(* Logix 5000 project; controller OWF Emulate 5570 rev 30.12; software revision 30.00; part 18 of 21 *)
(* tags used below, declared in another part *)
   OWF_Add_c : DINT;
   OWF_Input : DINT[16];
   OWF_Result : DINT[17];
(* MainProgram, continued *)

   		OWF_Result[4].31:=0;
   		OWF_Result[5]:=OWF_Result[5] + 1895099717+OWF_Add_c;
   		OWF_Add_c.5:=OWF_Result[5].31;
   		OWF_Result[5].31:=0;
   		OWF_Result[6]:=OWF_Result[6] + 2009701654+OWF_Add_c;
   		OWF_Add_c.6:=OWF_Result[6].31;
   		OWF_Result[6].31:=0;
   		OWF_Result[7]:=OWF_Result[7] + 1963030177+OWF_Add_c;
   		OWF_Add_c.7:=OWF_Result[7].31;
   		OWF_Result[7].31:=0;
   		OWF_Result[8]:=OWF_Result[8] + 232130595+OWF_Add_c;
   		OWF_Add_c.8:=OWF_Result[8].31;
   		OWF_Result[8].31:=0;
   		OWF_Result[9]:=OWF_Result[9] + 1484597708+OWF_Add_c;
   		OWF_Add_c.9:=OWF_Result[9].31;
   		OWF_Result[9].31:=0;
   		OWF_Result[10]:=OWF_Result[10] + 955822561+OWF_Add_c;
   		OWF_Add_c.10:=OWF_Result[10].31;
   		OWF_Result[10].31:=0;
   		OWF_Result[11]:=OWF_Result[11] + 760226904+OWF_Add_c;
   		OWF_Add_c.11:=OWF_Result[11].31;
   		OWF_Result[11].31:=0;
   		OWF_Result[12]:=OWF_Result[12] + 1637968730+OWF_Add_c;
   		OWF_Add_c.12:=OWF_Result[12].31;
   		OWF_Result[12].31:=0;
   		OWF_Result[13]:=OWF_Result[13] + 1060225387+OWF_Add_c;
   		OWF_Add_c.13:=OWF_Result[13].31;
   		OWF_Result[13].31:=0;
   		OWF_Result[14]:=OWF_Result[14] + 1695671309+OWF_Add_c;
   		OWF_Add_c.14:=OWF_Result[14].31;
   		OWF_Result[14].31:=0;
   		OWF_Result[15]:=OWF_Result[15] + 2141154184+OWF_Add_c;
   		OWF_Add_c.15:=OWF_Result[15].31;
   		OWF_Result[15].31:=0;
   		OWF_Result[16]:=OWF_Result[16] + 1403333060+OWF_Add_c;
   		OWF_Add_c.16:=OWF_Result[16].31;
   		OWF_Result[16].31:=0;
   	End_If;
   	If OWF_Input[11].[13] Then
   		OWF_Result[0]:=OWF_Result[0] + 1424989119+OWF_Add_c;
   		OWF_Add_c.0:=OWF_Result[0].31;
   		OWF_Result[0].31:=0;
   		OWF_Result[1]:=OWF_Result[1] + 1792831216+OWF_Add_c;
   		OWF_Add_c.1:=OWF_Result[1].31;
   		OWF_Result[1].31:=0;
   		OWF_Result[2]:=OWF_Result[2] + 1280480339+OWF_Add_c;
   		OWF_Add_c.2:=OWF_Result[2].31;
   		OWF_Result[2].31:=0;
   		OWF_Result[3]:=OWF_Result[3] + 1887620187+OWF_Add_c;
   		OWF_Add_c.3:=OWF_Result[3].31;
   		OWF_Result[3].31:=0;
   		OWF_Result[4]:=OWF_Result[4] + 50882950+OWF_Add_c;
   		OWF_Add_c.4:=OWF_Result[4].31;
   		OWF_Result[4].31:=0;
   		OWF_Result[5]:=OWF_Result[5] + 1542129432+OWF_Add_c;
   		OWF_Add_c.5:=OWF_Result[5].31;
   		OWF_Result[5].31:=0;
   		OWF_Result[6]:=OWF_Result[6] + 1234316724+OWF_Add_c;
   		OWF_Add_c.6:=OWF_Result[6].31;
   		OWF_Result[6].31:=0;
   		OWF_Result[7]:=OWF_Result[7] + 267891254+OWF_Add_c;
   		OWF_Add_c.7:=OWF_Result[7].31;
   		OWF_Result[7].31:=0;
   		OWF_Result[8]:=OWF_Result[8] + 1066053149+OWF_Add_c;
   		OWF_Add_c.8:=OWF_Result[8].31;
   		OWF_Result[8].31:=0;
   		OWF_Result[9]:=OWF_Result[9] + 54187296+OWF_Add_c;
   		OWF_Add_c.9:=OWF_Result[9].31;
   		OWF_Result[9].31:=0;
   		OWF_Result[10]:=OWF_Result[10] + 129651269+OWF_Add_c;
   		OWF_Add_c.10:=OWF_Result[10].31;
   		OWF_Result[10].31:=0;
   		OWF_Result[11]:=OWF_Result[11] + 604389954+OWF_Add_c;
   		OWF_Add_c.11:=OWF_Result[11].31;
   		OWF_Result[11].31:=0;
   		OWF_Result[12]:=OWF_Result[12] + 1474729667+OWF_Add_c;
   		OWF_Add_c.12:=OWF_Result[12].31;
   		OWF_Result[12].31:=0;
   		OWF_Result[13]:=OWF_Result[13] + 627513733+OWF_Add_c;
   		OWF_Add_c.13:=OWF_Result[13].31;
   		OWF_Result[13].31:=0;
   		OWF_Result[14]:=OWF_Result[14] + 1221285509+OWF_Add_c;
   		OWF_Add_c.14:=OWF_Result[14].31;
   		OWF_Result[14].31:=0;
   		OWF_Result[15]:=OWF_Result[15] + 1347886424+OWF_Add_c;
   		OWF_Add_c.15:=OWF_Result[15].31;
   		OWF_Result[15].31:=0;
   		OWF_Result[16]:=OWF_Result[16] + 1501741428+OWF_Add_c;
   		OWF_Add_c.16:=OWF_Result[16].31;
   		OWF_Result[16].31:=0;
   	End_If;
   	If OWF_Input[11].[14] Then
   		OWF_Result[0]:=OWF_Result[0] + 148251354+OWF_Add_c;
   		OWF_Add_c.0:=OWF_Result[0].31;
   		OWF_Result[0].31:=0;
   		OWF_Result[1]:=OWF_Result[1] + 734679875+OWF_Add_c;
   		OWF_Add_c.1:=OWF_Result[1].31;
   		OWF_Result[1].31:=0;
   		OWF_Result[2]:=OWF_Result[2] + 501019324+OWF_Add_c;
   		OWF_Add_c.2:=OWF_Result[2].31;
   		OWF_Result[2].31:=0;
   		OWF_Result[3]:=OWF_Result[3] + 1051894690+OWF_Add_c;
   		OWF_Add_c.3:=OWF_Result[3].31;
   		OWF_Result[3].31:=0;
   		OWF_Result[4]:=OWF_Result[4] + 713394787+OWF_Add_c;
   		OWF_Add_c.4:=OWF_Result[4].31;
   		OWF_Result[4].31:=0;
   		OWF_Result[5]:=OWF_Result[5] + 875122393+OWF_Add_c;
   		OWF_Add_c.5:=OWF_Result[5].31;
   		OWF_Result[5].31:=0;
   		OWF_Result[6]:=OWF_Result[6] + 259478417+OWF_Add_c;
   		OWF_Add_c.6:=OWF_Result[6].31;
   		OWF_Result[6].31:=0;
   		OWF_Result[7]:=OWF_Result[7] + 1855876414+OWF_Add_c;
   		OWF_Add_c.7:=OWF_Result[7].31;
   		OWF_Result[7].31:=0;
   		OWF_Result[8]:=OWF_Result[8] + 1892105+OWF_Add_c;
   		OWF_Add_c.8:=OWF_Result[8].31;
   		OWF_Result[8].31:=0;
   		OWF_Result[9]:=OWF_Result[9] + 229647947+OWF_Add_c;
   		OWF_Add_c.9:=OWF_Result[9].31;
   		OWF_Result[9].31:=0;
   		OWF_Result[10]:=OWF_Result[10] + 445153450+OWF_Add_c;
   		OWF_Add_c.10:=OWF_Result[10].31;
   		OWF_Result[10].31:=0;
   		OWF_Result[11]:=OWF_Result[11] + 1697696739+OWF_Add_c;
   		OWF_Add_c.11:=OWF_Result[11].31;
   		OWF_Result[11].31:=0;
   		OWF_Result[12]:=OWF_Result[12] + 259481221+OWF_Add_c;
   		OWF_Add_c.12:=OWF_Result[12].31;
   		OWF_Result[12].31:=0;
   		OWF_Result[13]:=OWF_Result[13] + 98481250+OWF_Add_c;
   		OWF_Add_c.13:=OWF_Result[13].31;
   		OWF_Result[13].31:=0;
   		OWF_Result[14]:=OWF_Result[14] + 6041701+OWF_Add_c;
   		OWF_Add_c.14:=OWF_Result[14].31;
   		OWF_Result[14].31:=0;
   		OWF_Result[15]:=OWF_Result[15] + 184524762+OWF_Add_c;
   		OWF_Add_c.15:=OWF_Result[15].31;
   		OWF_Result[15].31:=0;
   		OWF_Result[16]:=OWF_Result[16] + 729095478+OWF_Add_c;
   		OWF_Add_c.16:=OWF_Result[16].31;
   		OWF_Result[16].31:=0;
   	End_If;
   	If OWF_Input[11].[15] Then
   		OWF_Result[0]:=OWF_Result[0] + 681500769+OWF_Add_c;
   		OWF_Add_c.0:=OWF_Result[0].31;
   		OWF_Result[0].31:=0;
   		OWF_Result[1]:=OWF_Result[1] + 369563308+OWF_Add_c;
   		OWF_Add_c.1:=OWF_Result[1].31;
   		OWF_Result[1].31:=0;
   		OWF_Result[2]:=OWF_Result[2] + 577751378+OWF_Add_c;
   		OWF_Add_c.2:=OWF_Result[2].31;
   		OWF_Result[2].31:=0;
   		OWF_Result[3]:=OWF_Result[3] + 1178477344+OWF_Add_c;
   		OWF_Add_c.3:=OWF_Result[3].31;
   		OWF_Result[3].31:=0;
   		OWF_Result[4]:=OWF_Result[4] + 598929159+OWF_Add_c;
   		OWF_Add_c.4:=OWF_Result[4].31;
   		OWF_Result[4].31:=0;
   		OWF_Result[5]:=OWF_Result[5] + 1811347302+OWF_Add_c;
   		OWF_Add_c.5:=OWF_Result[5].31;
   		OWF_Result[5].31:=0;
   		OWF_Result[6]:=OWF_Result[6] + 309483525+OWF_Add_c;
   		OWF_Add_c.6:=OWF_Result[6].31;
   		OWF_Result[6].31:=0;
   		OWF_Result[7]:=OWF_Result[7] + 1944832940+OWF_Add_c;
   		OWF_Add_c.7:=OWF_Result[7].31;
   		OWF_Result[7].31:=0;
   		OWF_Result[8]:=OWF_Result[8] + 1640593669+OWF_Add_c;
   		OWF_Add_c.8:=OWF_Result[8].31;
   		OWF_Result[8].31:=0;
   		OWF_Result[9]:=OWF_Result[9] + 64106164+OWF_Add_c;
   		OWF_Add_c.9:=OWF_Result[9].31;
   		OWF_Result[9].31:=0;
   		OWF_Result[10]:=OWF_Result[10] + 1859760050+OWF_Add_c;
   		OWF_Add_c.10:=OWF_Result[10].31;
   		OWF_Result[10].31:=0;
   		OWF_Result[11]:=OWF_Result[11] + 1868576516+OWF_Add_c;
   		OWF_Add_c.11:=OWF_Result[11].31;
   		OWF_Result[11].31:=0;
   		OWF_Result[12]:=OWF_Result[12] + 1267284033+OWF_Add_c;
   		OWF_Add_c.12:=OWF_Result[12].31;
   		OWF_Result[12].31:=0;
   		OWF_Result[13]:=OWF_Result[13] + 1701199951+OWF_Add_c;
   		OWF_Add_c.13:=OWF_Result[13].31;
   		OWF_Result[13].31:=0;
   		OWF_Result[14]:=OWF_Result[14] + 2144306817+OWF_Add_c;
   		OWF_Add_c.14:=OWF_Result[14].31;
   		OWF_Result[14].31:=0;
   		OWF_Result[15]:=OWF_Result[15] + 1791762522+OWF_Add_c;
   		OWF_Add_c.15:=OWF_Result[15].31;
   		OWF_Result[15].31:=0;
   		OWF_Result[16]:=OWF_Result[16] + 81122948+OWF_Add_c;
   		OWF_Add_c.16:=OWF_Result[16].31;
   		OWF_Result[16].31:=0;
   	End_If;
   	If OWF_Input[11].[16] Then
   		OWF_Result[0]:=OWF_Result[0] + 17838217+OWF_Add_c;
   		OWF_Add_c.0:=OWF_Result[0].31;
   		OWF_Result[0].31:=0;
   		OWF_Result[1]:=OWF_Result[1] + 667401238+OWF_Add_c;
   		OWF_Add_c.1:=OWF_Result[1].31;
   		OWF_Result[1].31:=0;
   		OWF_Result[2]:=OWF_Result[2] + 325014797+OWF_Add_c;
   		OWF_Add_c.2:=OWF_Result[2].31;
   		OWF_Result[2].31:=0;
   		OWF_Result[3]:=OWF_Result[3] + 1946608283+OWF_Add_c;
   		OWF_Add_c.3:=OWF_Result[3].31;
   		OWF_Result[3].31:=0;
   		OWF_Result[4]:=OWF_Result[4] + 669694453+OWF_Add_c;
   		OWF_Add_c.4:=OWF_Result[4].31;
   		OWF_Result[4].31:=0;
   		OWF_Result[5]:=OWF_Result[5] + 261662885+OWF_Add_c;
   		OWF_Add_c.5:=OWF_Result[5].31;
   		OWF_Result[5].31:=0;
   		OWF_Result[6]:=OWF_Result[6] + 844241477+OWF_Add_c;
   		OWF_Add_c.6:=OWF_Result[6].31;
   		OWF_Result[6].31:=0;
   		OWF_Result[7]:=OWF_Result[7] + 1156660817+OWF_Add_c;
   		OWF_Add_c.7:=OWF_Result[7].31;
   		OWF_Result[7].31:=0;
   		OWF_Result[8]:=OWF_Result[8] + 1612944285+OWF_Add_c;
   		OWF_Add_c.8:=OWF_Result[8].31;
   		OWF_Result[8].31:=0;
   		OWF_Result[9]:=OWF_Result[9] + 1338738967+OWF_Add_c;
   		OWF_Add_c.9:=OWF_Result[9].31;
   		OWF_Result[9].31:=0;
   		OWF_Result[10]:=OWF_Result[10] + 1820634011+OWF_Add_c;
   		OWF_Add_c.10:=OWF_Result[10].31;
   		OWF_Result[10].31:=0;
   		OWF_Result[11]:=OWF_Result[11] + 612985796+OWF_Add_c;
   		OWF_Add_c.11:=OWF_Result[11].31;
   		OWF_Result[11].31:=0;
   		OWF_Result[12]:=OWF_Result[12] + 1546055205+OWF_Add_c;
   		OWF_Add_c.12:=OWF_Result[12].31;
   		OWF_Result[12].31:=0;
   		OWF_Result[13]:=OWF_Result[13] + 1420246016+OWF_Add_c;
   		OWF_Add_c.13:=OWF_Result[13].31;
   		OWF_Result[13].31:=0;
   		OWF_Result[14]:=OWF_Result[14] + 1971045595+OWF_Add_c;
   		OWF_Add_c.14:=OWF_Result[14].31;
   		OWF_Result[14].31:=0;
   		OWF_Result[15]:=OWF_Result[15] + 898490888+OWF_Add_c;
   		OWF_Add_c.15:=OWF_Result[15].31;
   		OWF_Result[15].31:=0;
   		OWF_Result[16]:=OWF_Result[16] + 301090578+OWF_Add_c;
   		OWF_Add_c.16:=OWF_Result[16].31;
   		OWF_Result[16].31:=0;
   	End_If;
   	If OWF_Input[11].[17] Then
   		OWF_Result[0]:=OWF_Result[0] + 1716459433+OWF_Add_c;
   		OWF_Add_c.0:=OWF_Result[0].31;
   		OWF_Result[0].31:=0;
   		OWF_Result[1]:=OWF_Result[1] + 50088708+OWF_Add_c;
   		OWF_Add_c.1:=OWF_Result[1].31;
   		OWF_Result[1].31:=0;
   		OWF_Result[2]:=OWF_Result[2] + 771574645+OWF_Add_c;
   		OWF_Add_c.2:=OWF_Result[2].31;
   		OWF_Result[2].31:=0;
   		OWF_Result[3]:=OWF_Result[3] + 141391603+OWF_Add_c;
   		OWF_Add_c.3:=OWF_Result[3].31;
   		OWF_Result[3].31:=0;
   		OWF_Result[4]:=OWF_Result[4] + 499486646+OWF_Add_c;
   		OWF_Add_c.4:=OWF_Result[4].31;
   		OWF_Result[4].31:=0;
   		OWF_Result[5]:=OWF_Result[5] + 1280378172+OWF_Add_c;
   		OWF_Add_c.5:=OWF_Result[5].31;
   		OWF_Result[5].31:=0;
   		OWF_Result[6]:=OWF_Result[6] + 205274223+OWF_Add_c;
   		OWF_Add_c.6:=OWF_Result[6].31;
   		OWF_Result[6].31:=0;
   		OWF_Result[7]:=OWF_Result[7] + 386848157+OWF_Add_c;
   		OWF_Add_c.7:=OWF_Result[7].31;
   		OWF_Result[7].31:=0;
   		OWF_Result[8]:=OWF_Result[8] + 1335980614+OWF_Add_c;
   		OWF_Add_c.8:=OWF_Result[8].31;
   		OWF_Result[8].31:=0;
   		OWF_Result[9]:=OWF_Result[9] + 1934630920+OWF_Add_c;
   		OWF_Add_c.9:=OWF_Result[9].31;
   		OWF_Result[9].31:=0;
   		OWF_Result[10]:=OWF_Result[10] + 271603978+OWF_Add_c;
   		OWF_Add_c.10:=OWF_Result[10].31;
   		OWF_Result[10].31:=0;
   		OWF_Result[11]:=OWF_Result[11] + 2088757329+OWF_Add_c;
   		OWF_Add_c.11:=OWF_Result[11].31;
   		OWF_Result[11].31:=0;
   		OWF_Result[12]:=OWF_Result[12] + 554669077+OWF_Add_c;
   		OWF_Add_c.12:=OWF_Result[12].31;
   		OWF_Result[12].31:=0;
   		OWF_Result[13]:=OWF_Result[13] + 1572623455+OWF_Add_c;
   		OWF_Add_c.13:=OWF_Result[13].31;
   		OWF_Result[13].31:=0;
   		OWF_Result[14]:=OWF_Result[14] + 1305661387+OWF_Add_c;
   		OWF_Add_c.14:=OWF_Result[14].31;
   		OWF_Result[14].31:=0;
   		OWF_Result[15]:=OWF_Result[15] + 1475736021+OWF_Add_c;
   		OWF_Add_c.15:=OWF_Result[15].31;
   		OWF_Result[15].31:=0;
   		OWF_Result[16]:=OWF_Result[16] + 761633792+OWF_Add_c;
   		OWF_Add_c.16:=OWF_Result[16].31;
   		OWF_Result[16].31:=0;
   	End_If;
   	If OWF_Input[11].[18] Then
   		OWF_Result[0]:=OWF_Result[0] + 1774213961+OWF_Add_c;
   		OWF_Add_c.0:=OWF_Result[0].31;
   		OWF_Result[0].31:=0;
   		OWF_Result[1]:=OWF_Result[1] + 1956173104+OWF_Add_c;
   		OWF_Add_c.1:=OWF_Result[1].31;
   		OWF_Result[1].31:=0;
   		OWF_Result[2]:=OWF_Result[2] + 370111830+OWF_Add_c;
   		OWF_Add_c.2:=OWF_Result[2].31;
   		OWF_Result[2].31:=0;
   		OWF_Result[3]:=OWF_Result[3] + 162529263+OWF_Add_c;
   		OWF_Add_c.3:=OWF_Result[3].31;
   		OWF_Result[3].31:=0;
   		OWF_Result[4]:=OWF_Result[4] + 2079589906+OWF_Add_c;
   		OWF_Add_c.4:=OWF_Result[4].31;
   		OWF_Result[4].31:=0;
   		OWF_Result[5]:=OWF_Result[5] + 725728807+OWF_Add_c;
   		OWF_Add_c.5:=OWF_Result[5].31;
   		OWF_Result[5].31:=0;
   		OWF_Result[6]:=OWF_Result[6] + 176946544+OWF_Add_c;
   		OWF_Add_c.6:=OWF_Result[6].31;
   		OWF_Result[6].31:=0;
   		OWF_Result[7]:=OWF_Result[7] + 1129912929+OWF_Add_c;
   		OWF_Add_c.7:=OWF_Result[7].31;
   		OWF_Result[7].31:=0;
   		OWF_Result[8]:=OWF_Result[8] + 1014363434+OWF_Add_c;
   		OWF_Add_c.8:=OWF_Result[8].31;
   		OWF_Result[8].31:=0;
   		OWF_Result[9]:=OWF_Result[9] + 1412304844+OWF_Add_c;
   		OWF_Add_c.9:=OWF_Result[9].31;
   		OWF_Result[9].31:=0;
   		OWF_Result[10]:=OWF_Result[10] + 141623841+OWF_Add_c;
   		OWF_Add_c.10:=OWF_Result[10].31;
   		OWF_Result[10].31:=0;
   		OWF_Result[11]:=OWF_Result[11] + 1305672224+OWF_Add_c;
   		OWF_Add_c.11:=OWF_Result[11].31;
   		OWF_Result[11].31:=0;
   		OWF_Result[12]:=OWF_Result[12] + 347830875+OWF_Add_c;
   		OWF_Add_c.12:=OWF_Result[12].31;
   		OWF_Result[12].31:=0;
   		OWF_Result[13]:=OWF_Result[13] + 1018422481+OWF_Add_c;
   		OWF_Add_c.13:=OWF_Result[13].31;
   		OWF_Result[13].31:=0;
   		OWF_Result[14]:=OWF_Result[14] + 1833122800+OWF_Add_c;
   		OWF_Add_c.14:=OWF_Result[14].31;
   		OWF_Result[14].31:=0;
   		OWF_Result[15]:=OWF_Result[15] + 1352323392+OWF_Add_c;
   		OWF_Add_c.15:=OWF_Result[15].31;
   		OWF_Result[15].31:=0;
   		OWF_Result[16]:=OWF_Result[16] + 490043194+OWF_Add_c;
   		OWF_Add_c.16:=OWF_Result[16].31;
   		OWF_Result[16].31:=0;
   	End_If;
   	If OWF_Input[11].[19] Then
   		OWF_Result[0]:=OWF_Result[0] + 1089958956+OWF_Add_c;
   		OWF_Add_c.0:=OWF_Result[0].31;
   		OWF_Result[0].31:=0;
   		OWF_Result[1]:=OWF_Result[1] + 147227708+OWF_Add_c;
   		OWF_Add_c.1:=OWF_Result[1].31;
   		OWF_Result[1].31:=0;
   		OWF_Result[2]:=OWF_Result[2] + 251643439+OWF_Add_c;
   		OWF_Add_c.2:=OWF_Result[2].31;
   		OWF_Result[2].31:=0;
   		OWF_Result[3]:=OWF_Result[3] + 1952477462+OWF_Add_c;
   		OWF_Add_c.3:=OWF_Result[3].31;
   		OWF_Result[3].31:=0;
   		OWF_Result[4]:=OWF_Result[4] + 752832647+OWF_Add_c;
   		OWF_Add_c.4:=OWF_Result[4].31;
   		OWF_Result[4].31:=0;
   		OWF_Result[5]:=OWF_Result[5] + 469694026+OWF_Add_c;
   		OWF_Add_c.5:=OWF_Result[5].31;
   		OWF_Result[5].31:=0;
   		OWF_Result[6]:=OWF_Result[6] + 84823545+OWF_Add_c;
   		OWF_Add_c.6:=OWF_Result[6].31;
   		OWF_Result[6].31:=0;
   		OWF_Result[7]:=OWF_Result[7] + 65062051+OWF_Add_c;
   		OWF_Add_c.7:=OWF_Result[7].31;
   		OWF_Result[7].31:=0;
   		OWF_Result[8]:=OWF_Result[8] + 2082323015+OWF_Add_c;
   		OWF_Add_c.8:=OWF_Result[8].31;
   		OWF_Result[8].31:=0;
   		OWF_Result[9]:=OWF_Result[9] + 1957541553+OWF_Add_c;
   		OWF_Add_c.9:=OWF_Result[9].31;
   		OWF_Result[9].31:=0;
   		OWF_Result[10]:=OWF_Result[10] + 881322145+OWF_Add_c;
   		OWF_Add_c.10:=OWF_Result[10].31;
   		OWF_Result[10].31:=0;
   		OWF_Result[11]:=OWF_Result[11] + 274678903+OWF_Add_c;
   		OWF_Add_c.11:=OWF_Result[11].31;
   		OWF_Result[11].31:=0;
   		OWF_Result[12]:=OWF_Result[12] + 2066464993+OWF_Add_c;
   		OWF_Add_c.12:=OWF_Result[12].31;
   		OWF_Result[12].31:=0;
   		OWF_Result[13]:=OWF_Result[13] + 1519945331+OWF_Add_c;
   		OWF_Add_c.13:=OWF_Result[13].31;
   		OWF_Result[13].31:=0;
   		OWF_Result[14]:=OWF_Result[14] + 1234570606+OWF_Add_c;
   		OWF_Add_c.14:=OWF_Result[14].31;
   		OWF_Result[14].31:=0;
   		OWF_Result[15]:=OWF_Result[15] + 727147104+OWF_Add_c;
   		OWF_Add_c.15:=OWF_Result[15].31;
   		OWF_Result[15].31:=0;
   		OWF_Result[16]:=OWF_Result[16] + 766198026+OWF_Add_c;
   		OWF_Add_c.16:=OWF_Result[16].31;
   		OWF_Result[16].31:=0;
   	End_If;
   	If OWF_Input[11].[20] Then
   		OWF_Result[0]:=OWF_Result[0] + 1364648256+OWF_Add_c;
   		OWF_Add_c.0:=OWF_Result[0].31;
   		OWF_Result[0].31:=0;
   		OWF_Result[1]:=OWF_Result[1] + 164927068+OWF_Add_c;
   		OWF_Add_c.1:=OWF_Result[1].31;
   		OWF_Result[1].31:=0;
   		OWF_Result[2]:=OWF_Result[2] + 937767971+OWF_Add_c;
   		OWF_Add_c.2:=OWF_Result[2].31;
   		OWF_Result[2].31:=0;
   		OWF_Result[3]:=OWF_Result[3] + 902258282+OWF_Add_c;
   		OWF_Add_c.3:=OWF_Result[3].31;
   		OWF_Result[3].31:=0;
   		OWF_Result[4]:=OWF_Result[4] + 800183826+OWF_Add_c;
   		OWF_Add_c.4:=OWF_Result[4].31;
   		OWF_Result[4].31:=0;
   		OWF_Result[5]:=OWF_Result[5] + 997138363+OWF_Add_c;
   		OWF_Add_c.5:=OWF_Result[5].31;
   		OWF_Result[5].31:=0;
   		OWF_Result[6]:=OWF_Result[6] + 1334209867+OWF_Add_c;
   		OWF_Add_c.6:=OWF_Result[6].31;
   		OWF_Result[6].31:=0;
   		OWF_Result[7]:=OWF_Result[7] + 13223971+OWF_Add_c;
   		OWF_Add_c.7:=OWF_Result[7].31;
   		OWF_Result[7].31:=0;
   		OWF_Result[8]:=OWF_Result[8] + 382532483+OWF_Add_c;
   		OWF_Add_c.8:=OWF_Result[8].31;
   		OWF_Result[8].31:=0;
   		OWF_Result[9]:=OWF_Result[9] + 2068009884+OWF_Add_c;
   		OWF_Add_c.9:=OWF_Result[9].31;
   		OWF_Result[9].31:=0;
   		OWF_Result[10]:=OWF_Result[10] + 956603858+OWF_Add_c;
   		OWF_Add_c.10:=OWF_Result[10].31;
   		OWF_Result[10].31:=0;
   		OWF_Result[11]:=OWF_Result[11] + 1536890465+OWF_Add_c;
   		OWF_Add_c.11:=OWF_Result[11].31;
   		OWF_Result[11].31:=0;
   		OWF_Result[12]:=OWF_Result[12] + 298774715+OWF_Add_c;
   		OWF_Add_c.12:=OWF_Result[12].31;
   		OWF_Result[12].31:=0;
   		OWF_Result[13]:=OWF_Result[13] + 2111597775+OWF_Add_c;
   		OWF_Add_c.13:=OWF_Result[13].31;
   		OWF_Result[13].31:=0;
   		OWF_Result[14]:=OWF_Result[14] + 2134082550+OWF_Add_c;
   		OWF_Add_c.14:=OWF_Result[14].31;
   		OWF_Result[14].31:=0;
   		OWF_Result[15]:=OWF_Result[15] + 951934122+OWF_Add_c;
   		OWF_Add_c.15:=OWF_Result[15].31;
   		OWF_Result[15].31:=0;
   		OWF_Result[16]:=OWF_Result[16] + 443405783+OWF_Add_c;
   		OWF_Add_c.16:=OWF_Result[16].31;
   		OWF_Result[16].31:=0;
   	End_If;
   	If OWF_Input[11].[21] Then
   		OWF_Result[0]:=OWF_Result[0] + 1626999370+OWF_Add_c;
   		OWF_Add_c.0:=OWF_Result[0].31;
   		OWF_Result[0].31:=0;
   		OWF_Result[1]:=OWF_Result[1] + 563410518+OWF_Add_c;
   		OWF_Add_c.1:=OWF_Result[1].31;
   		OWF_Result[1].31:=0;
   		OWF_Result[2]:=OWF_Result[2] + 448996783+OWF_Add_c;
   		OWF_Add_c.2:=OWF_Result[2].31;
   		OWF_Result[2].31:=0;
   		OWF_Result[3]:=OWF_Result[3] + 1482249525+OWF_Add_c;
   		OWF_Add_c.3:=OWF_Result[3].31;
   		OWF_Result[3].31:=0;
   		OWF_Result[4]:=OWF_Result[4] + 1968681288+OWF_Add_c;
   		OWF_Add_c.4:=OWF_Result[4].31;
   		OWF_Result[4].31:=0;
   		OWF_Result[5]:=OWF_Result[5] + 289272502+OWF_Add_c;
   		OWF_Add_c.5:=OWF_Result[5].31;
   		OWF_Result[5].31:=0;
   		OWF_Result[6]:=OWF_Result[6] + 622481402+OWF_Add_c;
   		OWF_Add_c.6:=OWF_Result[6].31;
   		OWF_Result[6].31:=0;
   		OWF_Result[7]:=OWF_Result[7] + 1182960437+OWF_Add_c;
   		OWF_Add_c.7:=OWF_Result[7].31;
   		OWF_Result[7].31:=0;
   		OWF_Result[8]:=OWF_Result[8] + 194816774+OWF_Add_c;
   		OWF_Add_c.8:=OWF_Result[8].31;
   		OWF_Result[8].31:=0;
   		OWF_Result[9]:=OWF_Result[9] + 179922716+OWF_Add_c;
   		OWF_Add_c.9:=OWF_Result[9].31;
   		OWF_Result[9].31:=0;
   		OWF_Result[10]:=OWF_Result[10] + 393221600+OWF_Add_c;
   		OWF_Add_c.10:=OWF_Result[10].31;
   		OWF_Result[10].31:=0;
   		OWF_Result[11]:=OWF_Result[11] + 521638735+OWF_Add_c;
   		OWF_Add_c.11:=OWF_Result[11].31;
   		OWF_Result[11].31:=0;
   		OWF_Result[12]:=OWF_Result[12] + 1901625421+OWF_Add_c;
   		OWF_Add_c.12:=OWF_Result[12].31;
   		OWF_Result[12].31:=0;
   		OWF_Result[13]:=OWF_Result[13] + 1059351231+OWF_Add_c;
   		OWF_Add_c.13:=OWF_Result[13].31;
   		OWF_Result[13].31:=0;
   		OWF_Result[14]:=OWF_Result[14] + 133998538+OWF_Add_c;
   		OWF_Add_c.14:=OWF_Result[14].31;
   		OWF_Result[14].31:=0;
   		OWF_Result[15]:=OWF_Result[15] + 336969007+OWF_Add_c;
   		OWF_Add_c.15:=OWF_Result[15].31;
   		OWF_Result[15].31:=0;
   		OWF_Result[16]:=OWF_Result[16] + 1951770492+OWF_Add_c;
   		OWF_Add_c.16:=OWF_Result[16].31;
   		OWF_Result[16].31:=0;
   	End_If;
   	If OWF_Input[11].[22] Then
   		OWF_Result[0]:=OWF_Result[0] + 894773317+OWF_Add_c;
   		OWF_Add_c.0:=OWF_Result[0].31;
   		OWF_Result[0].31:=0;
   		OWF_Result[1]:=OWF_Result[1] + 606366330+OWF_Add_c;
   		OWF_Add_c.1:=OWF_Result[1].31;
   		OWF_Result[1].31:=0;
   		OWF_Result[2]:=OWF_Result[2] + 317214561+OWF_Add_c;
   		OWF_Add_c.2:=OWF_Result[2].31;
   		OWF_Result[2].31:=0;
   		OWF_Result[3]:=OWF_Result[3] + 1260101015+OWF_Add_c;
   		OWF_Add_c.3:=OWF_Result[3].31;
   		OWF_Result[3].31:=0;
   		OWF_Result[4]:=OWF_Result[4] + 1318837221+OWF_Add_c;
   		OWF_Add_c.4:=OWF_Result[4].31;
   		OWF_Result[4].31:=0;
   		OWF_Result[5]:=OWF_Result[5] + 301123999+OWF_Add_c;
   		OWF_Add_c.5:=OWF_Result[5].31;
   		OWF_Result[5].31:=0;
   		OWF_Result[6]:=OWF_Result[6] + 1904419438+OWF_Add_c;
   		OWF_Add_c.6:=OWF_Result[6].31;
   		OWF_Result[6].31:=0;
   		OWF_Result[7]:=OWF_Result[7] + 1567980401+OWF_Add_c;
   		OWF_Add_c.7:=OWF_Result[7].31;
   		OWF_Result[7].31:=0;
   		OWF_Result[8]:=OWF_Result[8] + 1450680308+OWF_Add_c;
   		OWF_Add_c.8:=OWF_Result[8].31;
   		OWF_Result[8].31:=0;
   		OWF_Result[9]:=OWF_Result[9] + 2141190341+OWF_Add_c;
   		OWF_Add_c.9:=OWF_Result[9].31;
   		OWF_Result[9].31:=0;
   		OWF_Result[10]:=OWF_Result[10] + 1361621893+OWF_Add_c;
   		OWF_Add_c.10:=OWF_Result[10].31;
   		OWF_Result[10].31:=0;
   		OWF_Result[11]:=OWF_Result[11] + 522285678+OWF_Add_c;
   		OWF_Add_c.11:=OWF_Result[11].31;
   		OWF_Result[11].31:=0;
   		OWF_Result[12]:=OWF_Result[12] + 1292342478+OWF_Add_c;
   		OWF_Add_c.12:=OWF_Result[12].31;
   		OWF_Result[12].31:=0;
   		OWF_Result[13]:=OWF_Result[13] + 1573930208+OWF_Add_c;
   		OWF_Add_c.13:=OWF_Result[13].31;
   		OWF_Result[13].31:=0;
   		OWF_Result[14]:=OWF_Result[14] + 578592603+OWF_Add_c;
   		OWF_Add_c.14:=OWF_Result[14].31;
   		OWF_Result[14].31:=0;
   		OWF_Result[15]:=OWF_Result[15] + 1531371679+OWF_Add_c;
   		OWF_Add_c.15:=OWF_Result[15].31;
   		OWF_Result[15].31:=0;
   		OWF_Result[16]:=OWF_Result[16] + 1500250328+OWF_Add_c;
   		OWF_Add_c.16:=OWF_Result[16].31;
   		OWF_Result[16].31:=0;
   	End_If;
   	If OWF_Input[11].[23] Then
   		OWF_Result[0]:=OWF_Result[0] + 1886057312+OWF_Add_c;
   		OWF_Add_c.0:=OWF_Result[0].31;
   		OWF_Result[0].31:=0;
   		OWF_Result[1]:=OWF_Result[1] + 1273986779+OWF_Add_c;
   		OWF_Add_c.1:=OWF_Result[1].31;
   		OWF_Result[1].31:=0;
   		OWF_Result[2]:=OWF_Result[2] + 1832540527+OWF_Add_c;
   		OWF_Add_c.2:=OWF_Result[2].31;
   		OWF_Result[2].31:=0;
   		OWF_Result[3]:=OWF_Result[3] + 1904028625+OWF_Add_c;
   		OWF_Add_c.3:=OWF_Result[3].31;
   		OWF_Result[3].31:=0;
   		OWF_Result[4]:=OWF_Result[4] + 166664105+OWF_Add_c;
   		OWF_Add_c.4:=OWF_Result[4].31;
   		OWF_Result[4].31:=0;
   		OWF_Result[5]:=OWF_Result[5] + 461900417+OWF_Add_c;
   		OWF_Add_c.5:=OWF_Result[5].31;
   		OWF_Result[5].31:=0;
   		OWF_Result[6]:=OWF_Result[6] + 1086720032+OWF_Add_c;
   		OWF_Add_c.6:=OWF_Result[6].31;
   		OWF_Result[6].31:=0;
   		OWF_Result[7]:=OWF_Result[7] + 1409617277+OWF_Add_c;
   		OWF_Add_c.7:=OWF_Result[7].31;
   		OWF_Result[7].31:=0;
   		OWF_Result[8]:=OWF_Result[8] + 391672452+OWF_Add_c;
   		OWF_Add_c.8:=OWF_Result[8].31;
   		OWF_Result[8].31:=0;
   		OWF_Result[9]:=OWF_Result[9] + 248948740+OWF_Add_c;
   		OWF_Add_c.9:=OWF_Result[9].31;
   		OWF_Result[9].31:=0;
   		OWF_Result[10]:=OWF_Result[10] + 767259363+OWF_Add_c;
   		OWF_Add_c.10:=OWF_Result[10].31;
   		OWF_Result[10].31:=0;
   		OWF_Result[11]:=OWF_Result[11] + 1785063648+OWF_Add_c;
   		OWF_Add_c.11:=OWF_Result[11].31;
   		OWF_Result[11].31:=0;
   		OWF_Result[12]:=OWF_Result[12] + 1895212709+OWF_Add_c;
   		OWF_Add_c.12:=OWF_Result[12].31;
   		OWF_Result[12].31:=0;
   		OWF_Result[13]:=OWF_Result[13] + 403462174+OWF_Add_c;
   		OWF_Add_c.13:=OWF_Result[13].31;
   		OWF_Result[13].31:=0;
   		OWF_Result[14]:=OWF_Result[14] + 1785074148+OWF_Add_c;
   		OWF_Add_c.14:=OWF_Result[14].31;
   		OWF_Result[14].31:=0;
   		OWF_Result[15]:=OWF_Result[15] + 1011949593+OWF_Add_c;
   		OWF_Add_c.15:=OWF_Result[15].31;
   		OWF_Result[15].31:=0;
   		OWF_Result[16]:=OWF_Result[16] + 1210282205+OWF_Add_c;
   		OWF_Add_c.16:=OWF_Result[16].31;
   		OWF_Result[16].31:=0;
   	End_If;
   	If OWF_Input[11].[24] Then
   		OWF_Result[0]:=OWF_Result[0] + 401282675+OWF_Add_c;
   		OWF_Add_c.0:=OWF_Result[0].31;
   		OWF_Result[0].31:=0;
   		OWF_Result[1]:=OWF_Result[1] + 799238946+OWF_Add_c;
   		OWF_Add_c.1:=OWF_Result[1].31;
   		OWF_Result[1].31:=0;
   		OWF_Result[2]:=OWF_Result[2] + 986211483+OWF_Add_c;
   		OWF_Add_c.2:=OWF_Result[2].31;
   		OWF_Result[2].31:=0;
   		OWF_Result[3]:=OWF_Result[3] + 934076381+OWF_Add_c;
   		OWF_Add_c.3:=OWF_Result[3].31;
   		OWF_Result[3].31:=0;
   		OWF_Result[4]:=OWF_Result[4] + 1371917488+OWF_Add_c;
   		OWF_Add_c.4:=OWF_Result[4].31;
   		OWF_Result[4].31:=0;
   		OWF_Result[5]:=OWF_Result[5] + 825496883+OWF_Add_c;
   		OWF_Add_c.5:=OWF_Result[5].31;
   		OWF_Result[5].31:=0;
   		OWF_Result[6]:=OWF_Result[6] + 1614904684+OWF_Add_c;
   		OWF_Add_c.6:=OWF_Result[6].31;
   		OWF_Result[6].31:=0;
   		OWF_Result[7]:=OWF_Result[7] + 801924968+OWF_Add_c;
   		OWF_Add_c.7:=OWF_Result[7].31;
   		OWF_Result[7].31:=0;
   		OWF_Result[8]:=OWF_Result[8] + 1059572265+OWF_Add_c;
   		OWF_Add_c.8:=OWF_Result[8].31;
   		OWF_Result[8].31:=0;
   		OWF_Result[9]:=OWF_Result[9] + 904716320+OWF_Add_c;
   		OWF_Add_c.9:=OWF_Result[9].31;
   		OWF_Result[9].31:=0;
   		OWF_Result[10]:=OWF_Result[10] + 1107544875+OWF_Add_c;
   		OWF_Add_c.10:=OWF_Result[10].31;
   		OWF_Result[10].31:=0;
   		OWF_Result[11]:=OWF_Result[11] + 1879948129+OWF_Add_c;
   		OWF_Add_c.11:=OWF_Result[11].31;
   		OWF_Result[11].31:=0;
   		OWF_Result[12]:=OWF_Result[12] + 1939277562+OWF_Add_c;
   		OWF_Add_c.12:=OWF_Result[12].31;
   		OWF_Result[12].31:=0;
   		OWF_Result[13]:=OWF_Result[13] + 1525082456+OWF_Add_c;
   		OWF_Add_c.13:=OWF_Result[13].31;
   		OWF_Result[13].31:=0;
   		OWF_Result[14]:=OWF_Result[14] + 1211143029+OWF_Add_c;
   		OWF_Add_c.14:=OWF_Result[14].31;
   		OWF_Result[14].31:=0;
   		OWF_Result[15]:=OWF_Result[15] + 1300216374+OWF_Add_c;
   		OWF_Add_c.15:=OWF_Result[15].31;
   		OWF_Result[15].31:=0;
   		OWF_Result[16]:=OWF_Result[16] + 1313625189+OWF_Add_c;
   		OWF_Add_c.16:=OWF_Result[16].31;
   		OWF_Result[16].31:=0;
   	End_If;
   	If OWF_Input[11].[25] Then
   		OWF_Result[0]:=OWF_Result[0] + 1056361843+OWF_Add_c;
   		OWF_Add_c.0:=OWF_Result[0].31;
   		OWF_Result[0].31:=0;
   		OWF_Result[1]:=OWF_Result[1] + 345909521+OWF_Add_c;
   		OWF_Add_c.1:=OWF_Result[1].31;
   		OWF_Result[1].31:=0;
   		OWF_Result[2]:=OWF_Result[2] + 1780659920+OWF_Add_c;
   		OWF_Add_c.2:=OWF_Result[2].31;
   		OWF_Result[2].31:=0;
   		OWF_Result[3]:=OWF_Result[3] + 1122260984+OWF_Add_c;
   		OWF_Add_c.3:=OWF_Result[3].31;
   		OWF_Result[3].31:=0;
   		OWF_Result[4]:=OWF_Result[4] + 1782435452+OWF_Add_c;
   		OWF_Add_c.4:=OWF_Result[4].31;
   		OWF_Result[4].31:=0;
   		OWF_Result[5]:=OWF_Result[5] + 1252964796+OWF_Add_c;
   		OWF_Add_c.5:=OWF_Result[5].31;
   		OWF_Result[5].31:=0;
   		OWF_Result[6]:=OWF_Result[6] + 1907967606+OWF_Add_c;
   		OWF_Add_c.6:=OWF_Result[6].31;
   		OWF_Result[6].31:=0;
   		OWF_Result[7]:=OWF_Result[7] + 906297812+OWF_Add_c;
   		OWF_Add_c.7:=OWF_Result[7].31;
   		OWF_Result[7].31:=0;
   		OWF_Result[8]:=OWF_Result[8] + 683910837+OWF_Add_c;
   		OWF_Add_c.8:=OWF_Result[8].31;
   		OWF_Result[8].31:=0;
   		OWF_Result[9]:=OWF_Result[9] + 1193260594+OWF_Add_c;
   		OWF_Add_c.9:=OWF_Result[9].31;
   		OWF_Result[9].31:=0;
   		OWF_Result[10]:=OWF_Result[10] + 958800894+OWF_Add_c;
   		OWF_Add_c.10:=OWF_Result[10].31;
   		OWF_Result[10].31:=0;
   		OWF_Result[11]:=OWF_Result[11] + 2018856363+OWF_Add_c;
   		OWF_Add_c.11:=OWF_Result[11].31;
   		OWF_Result[11].31:=0;
   		OWF_Result[12]:=OWF_Result[12] + 1253997947+OWF_Add_c;
   		OWF_Add_c.12:=OWF_Result[12].31;
   		OWF_Result[12].31:=0;
   		OWF_Result[13]:=OWF_Result[13] + 1085374324+OWF_Add_c;
   		OWF_Add_c.13:=OWF_Result[13].31;
   		OWF_Result[13].31:=0;
   		OWF_Result[14]:=OWF_Result[14] + 1969678640+OWF_Add_c;
   		OWF_Add_c.14:=OWF_Result[14].31;
   		OWF_Result[14].31:=0;
   		OWF_Result[15]:=OWF_Result[15] + 1714708581+OWF_Add_c;
   		OWF_Add_c.15:=OWF_Result[15].31;
   		OWF_Result[15].31:=0;
   		OWF_Result[16]:=OWF_Result[16] + 427066529+OWF_Add_c;
   		OWF_Add_c.16:=OWF_Result[16].31;
   		OWF_Result[16].31:=0;
   	End_If;
   	If OWF_Input[11].[26] Then
   		OWF_Result[0]:=OWF_Result[0] + 1013673849+OWF_Add_c;
   		OWF_Add_c.0:=OWF_Result[0].31;
   		OWF_Result[0].31:=0;
   		OWF_Result[1]:=OWF_Result[1] + 599971454+OWF_Add_c;
   		OWF_Add_c.1:=OWF_Result[1].31;
   		OWF_Result[1].31:=0;
   		OWF_Result[2]:=OWF_Result[2] + 644478275+OWF_Add_c;
   		OWF_Add_c.2:=OWF_Result[2].31;
   		OWF_Result[2].31:=0;
   		OWF_Result[3]:=OWF_Result[3] + 1083158658+OWF_Add_c;
   		OWF_Add_c.3:=OWF_Result[3].31;
   		OWF_Result[3].31:=0;
   		OWF_Result[4]:=OWF_Result[4] + 259583700+OWF_Add_c;
   		OWF_Add_c.4:=OWF_Result[4].31;
   		OWF_Result[4].31:=0;
   		OWF_Result[5]:=OWF_Result[5] + 61386803+OWF_Add_c;
   		OWF_Add_c.5:=OWF_Result[5].31;
   		OWF_Result[5].31:=0;
   		OWF_Result[6]:=OWF_Result[6] + 242575109+OWF_Add_c;
   		OWF_Add_c.6:=OWF_Result[6].31;
   		OWF_Result[6].31:=0;
   		OWF_Result[7]:=OWF_Result[7] + 1595828400+OWF_Add_c;
   		OWF_Add_c.7:=OWF_Result[7].31;
   		OWF_Result[7].31:=0;
   		OWF_Result[8]:=OWF_Result[8] + 1472352741+OWF_Add_c;
   		OWF_Add_c.8:=OWF_Result[8].31;
   		OWF_Result[8].31:=0;
   		OWF_Result[9]:=OWF_Result[9] + 2137321336+OWF_Add_c;
   		OWF_Add_c.9:=OWF_Result[9].31;
   		OWF_Result[9].31:=0;
   		OWF_Result[10]:=OWF_Result[10] + 670771411+OWF_Add_c;
   		OWF_Add_c.10:=OWF_Result[10].31;
   		OWF_Result[10].31:=0;
   		OWF_Result[11]:=OWF_Result[11] + 1778817064+OWF_Add_c;
   		OWF_Add_c.11:=OWF_Result[11].31;
   		OWF_Result[11].31:=0;
   		OWF_Result[12]:=OWF_Result[12] + 1118459420+OWF_Add_c;
   		OWF_Add_c.12:=OWF_Result[12].31;
   		OWF_Result[12].31:=0;
   		OWF_Result[13]:=OWF_Result[13] + 892634991+OWF_Add_c;
   		OWF_Add_c.13:=OWF_Result[13].31;
   		OWF_Result[13].31:=0;
   		OWF_Result[14]:=OWF_Result[14] + 775096057+OWF_Add_c;
   		OWF_Add_c.14:=OWF_Result[14].31;
   		OWF_Result[14].31:=0;
   		OWF_Result[15]:=OWF_Result[15] + 1710450555+OWF_Add_c;
   		OWF_Add_c.15:=OWF_Result[15].31;
   		OWF_Result[15].31:=0;
   		OWF_Result[16]:=OWF_Result[16] + 1568308360+OWF_Add_c;
   		OWF_Add_c.16:=OWF_Result[16].31;
   		OWF_Result[16].31:=0;
   	End_If;
   	If OWF_Input[11].[27] Then
   		OWF_Result[0]:=OWF_Result[0] + 66795224+OWF_Add_c;
   		OWF_Add_c.0:=OWF_Result[0].31;
   		OWF_Result[0].31:=0;
   		OWF_Result[1]:=OWF_Result[1] + 1940340644+OWF_Add_c;
   		OWF_Add_c.1:=OWF_Result[1].31;
   		OWF_Result[1].31:=0;
   		OWF_Result[2]:=OWF_Result[2] + 631847958+OWF_Add_c;
   		OWF_Add_c.2:=OWF_Result[2].31;
   		OWF_Result[2].31:=0;
   		OWF_Result[3]:=OWF_Result[3] + 427458976+OWF_Add_c;
   		OWF_Add_c.3:=OWF_Result[3].31;
   		OWF_Result[3].31:=0;
   		OWF_Result[4]:=OWF_Result[4] + 1873358097+OWF_Add_c;
   		OWF_Add_c.4:=OWF_Result[4].31;
   		OWF_Result[4].31:=0;
   		OWF_Result[5]:=OWF_Result[5] + 1298619133+OWF_Add_c;
   		OWF_Add_c.5:=OWF_Result[5].31;
   		OWF_Result[5].31:=0;
   		OWF_Result[6]:=OWF_Result[6] + 849957863+OWF_Add_c;
   		OWF_Add_c.6:=OWF_Result[6].31;
   		OWF_Result[6].31:=0;
   		OWF_Result[7]:=OWF_Result[7] + 342461804+OWF_Add_c;
   		OWF_Add_c.7:=OWF_Result[7].31;
   		OWF_Result[7].31:=0;
   		OWF_Result[8]:=OWF_Result[8] + 458536952+OWF_Add_c;
   		OWF_Add_c.8:=OWF_Result[8].31;
   		OWF_Result[8].31:=0;
   		OWF_Result[9]:=OWF_Result[9] + 991963534+OWF_Add_c;
   		OWF_Add_c.9:=OWF_Result[9].31;
   		OWF_Result[9].31:=0;
   		OWF_Result[10]:=OWF_Result[10] + 374452693+OWF_Add_c;
   		OWF_Add_c.10:=OWF_Result[10].31;
   		OWF_Result[10].31:=0;
   		OWF_Result[11]:=OWF_Result[11] + 24063952+OWF_Add_c;
   		OWF_Add_c.11:=OWF_Result[11].31;
   		OWF_Result[11].31:=0;
   		OWF_Result[12]:=OWF_Result[12] + 1826661064+OWF_Add_c;
   		OWF_Add_c.12:=OWF_Result[12].31;
   		OWF_Result[12].31:=0;
   		OWF_Result[13]:=OWF_Result[13] + 23293515+OWF_Add_c;
   		OWF_Add_c.13:=OWF_Result[13].31;
   		OWF_Result[13].31:=0;
   		OWF_Result[14]:=OWF_Result[14] + 1732775983+OWF_Add_c;
   		OWF_Add_c.14:=OWF_Result[14].31;